   TS[126].ALLG.POS.End_1 := 491999;
   TS[126].ALLG.Stop_Position := 7200;
   TS[126].ALLG.Drive_speed_1 := 15000;
   TS[126].ALLG.Drive_speed_2 := 10000;
   TS[127].ALLG.POS.Start_1 := 492000;
   TS[127].ALLG.POS.End_1 := 498199;
   TS[127].ALLG.Stop_Position := 5400;
   TS[127].ALLG.Drive_speed_1 := 15000;
   TS[127].ALLG.Drive_speed_2 := 10000;
   TS[128].ALLG.POS.Start_1 := 498200;
   TS[128].ALLG.POS.End_1 := 504399;
   TS[128].ALLG.Stop_Position := 2954;
   TS[128].ALLG.Drive_speed_1 := 15000;
   TS[128].ALLG.Drive_speed_2 := 10000;
   TS[129].ALLG.POS.Start_1 := 504400;
   TS[129].ALLG.POS.End_1 := 511399;
   TS[129].ALLG.Stop_Position := 6300;
   TS[129].ALLG.Drive_speed_1 := 15000;
   TS[129].ALLG.Drive_speed_2 := 10000;
   TS[130].ALLG.POS.Start_1 := 511400;
   TS[130].ALLG.POS.End_1 := 518399;
   TS[130].ALLG.Stop_Position := 6300;
   TS[130].ALLG.Drive_speed_1 := 15000;
   TS[130].ALLG.Drive_speed_2 := 10000;
   TS[131].ALLG.POS.Start_1 := 518400;
   TS[131].ALLG.POS.End_1 := 525599;
   TS[131].ALLG.Stop_Position := 6300;
   TS[131].ALLG.Drive_speed_1 := 15000;
   TS[131].ALLG.Drive_speed_2 := 10000;
   TS[132].ALLG.POS.Start_1 := 525600;
   TS[132].ALLG.POS.End_1 := 529699;
   TS[132].ALLG.Stop_Position := 4299;
   TS[132].ALLG.Drive_speed_1 := 10000;
   TS[132].ALLG.Drive_speed_2 := 10000;
   TS[140].ALLG.POS.Start_1 := 529700;
   TS[140].ALLG.POS.End_1 := 535699;
   TS[140].ALLG.Stop_Position := 5900;
   TS[140].ALLG.Drive_speed_1 := 30000;
   TS[140].ALLG.Drive_speed_2 := 10000;
   TS[141].ALLG.POS.Start_1 := 535700;
   TS[141].ALLG.POS.End_1 := 541699;
   TS[141].ALLG.Stop_Position := 5900;
   TS[141].ALLG.Drive_speed_1 := 30000;
   TS[141].ALLG.Drive_speed_2 := 10000;
   TS[142].ALLG.POS.Start_1 := 541700;
   TS[142].ALLG.POS.End_1 := 547699;
   TS[142].ALLG.Stop_Position := 5900;
   TS[142].ALLG.Drive_speed_1 := 30000;
   TS[142].ALLG.Drive_speed_2 := 10000;
   TS[143].ALLG.POS.Start_1 := 547700;
   TS[143].ALLG.POS.End_1 := 553699;
   TS[143].ALLG.Stop_Position := 5900;
   TS[143].ALLG.Drive_speed_1 := 30000;
   TS[143].ALLG.Drive_speed_2 := 10000;
   TS[144].ALLG.POS.Start_1 := 553700;
   TS[144].ALLG.POS.End_1 := 559699;
   TS[144].ALLG.Stop_Position := 5900;
   TS[144].ALLG.Drive_speed_1 := 30000;
   TS[144].ALLG.Drive_speed_2 := 10000;
   TS[145].ALLG.POS.Start_1 := 559700;
   TS[145].ALLG.POS.End_1 := 565699;
   TS[145].ALLG.Stop_Position := 5900;
   TS[145].ALLG.Drive_speed_1 := 30000;
   TS[145].ALLG.Drive_speed_2 := 10000;
   TS[146].ALLG.POS.Start_1 := 565700;
   TS[146].ALLG.POS.End_1 := 571699;
   TS[146].ALLG.Stop_Position := 5900;
   TS[146].ALLG.Drive_speed_1 := 30000;
   TS[146].ALLG.Drive_speed_2 := 10000;
   TS[147].ALLG.POS.Start_1 := 571700;
   TS[147].ALLG.POS.End_1 := 577699;
   TS[147].ALLG.Stop_Position := 5900;
   TS[147].ALLG.Drive_speed_1 := 30000;
   TS[147].ALLG.Drive_speed_2 := 10000;
   TS[148].ALLG.POS.Start_1 := 577700;
   TS[148].ALLG.POS.End_1 := 583699;
   TS[148].ALLG.Stop_Position := 5900;
   TS[148].ALLG.Drive_speed_1 := 30000;
   TS[148].ALLG.Drive_speed_2 := 10000;
   TS[149].ALLG.POS.Start_1 := 583700;
   TS[149].ALLG.POS.End_1 := 589699;
   TS[149].ALLG.Stop_Position := 5900;
   TS[149].ALLG.Drive_speed_1 := 30000;
   TS[149].ALLG.Drive_speed_2 := 10000;
   TS[150].ALLG.POS.Start_1 := 589700;
   TS[150].ALLG.POS.End_1 := 595699;
   TS[150].ALLG.Stop_Position := 5900;
   TS[150].ALLG.Drive_speed_1 := 25000;
   TS[150].ALLG.Drive_speed_2 := 10000;
   TS[151].ALLG.POS.Start_1 := 595700;
   TS[151].ALLG.POS.End_1 := 601699;
   TS[151].ALLG.Stop_Position := 5900;
   TS[151].ALLG.Drive_speed_1 := 18000;
   TS[151].ALLG.Drive_speed_2 := 10000;
   TS[152].ALLG.POS.Start_1 := 601700;
   TS[152].ALLG.POS.End_1 := 607699;
   TS[152].ALLG.Stop_Position := 5900;
   TS[152].ALLG.Drive_speed_1 := 18000;
   TS[152].ALLG.Drive_speed_2 := 10000;
   TS[160].ALLG.POS.Start_1 := 607700;
   TS[160].ALLG.POS.End_1 := 613699;
   TS[160].ALLG.Stop_Position := 5900;
   TS[160].ALLG.Drive_speed_1 := 20000;
   TS[160].ALLG.Drive_speed_2 := 10000;
   TS[161].ALLG.POS.Start_1 := 613700;
   TS[161].ALLG.POS.End_1 := 619699;
   TS[161].ALLG.Stop_Position := 5900;
   TS[161].ALLG.Drive_speed_1 := 20000;
   TS[161].ALLG.Drive_speed_2 := 10000;
   TS[162].ALLG.POS.Start_1 := 619700;
   TS[162].ALLG.POS.End_1 := 625699;
   TS[162].ALLG.Stop_Position := 5900;
   TS[162].ALLG.Drive_speed_1 := 20000;
   TS[162].ALLG.Drive_speed_2 := 10000;
   // 15300 more start values not shown
END_DATA_BLOCK

DATA_BLOCK "DB_SDC_TS_PARAMETER_3"   // DB3706
{ S7_Optimized_Access := 'FALSE' }
AUTHOR : FFM
FAMILY : SDC
NAME : SECT_DEF
VERSION : 1.0
   VAR
      HEADER : Struct   // Struktur für Datenheader // nicht verschieben
         DB_NR : Int := 3706;   // DB Nummer
         MIN_NR_SEK : Int := 201;   // Niedrigste SEK Nummer im DB
         MAX_NR_SEK : Int := 300;   // Höchste SEK Nummer im DB
         START_DAT : Int := 20;   // Startadresse der SEK im DB
         LAENGE_SEK_DATA : Int := 260;   // Länge SEK Data
         ANZ_PROFIL : Int := 10;   // Number of Profiles
         OFFEST_PROFIL : Int := 40;   // Offestadresse der Profilparameter im TS-Parameterdatensatz
         LAENGE_PROFIL_DATA : Int := 22;   // Länge SEK Data
         Res160 : Int := 0;   // Reserve
         Res : Int := 0;   // Reserve
      END_STRUCT;
      TS : Array[201..300] of "UDT_SDC_TS_PARAMETER";
   END_VAR
BEGIN
   TS[201].ALLG.SEK_NEXT_1 := 0;
   TS[201].ALLG.SEK_NEXT_2 := 0;
   TS[201].ALLG.Spare[4] := 16#00;
   TS[201].ALLG.Spare[5] := 16#00;
   TS[201].ALLG.POS.Start_1 := 709550;
   TS[201].ALLG.POS.End_1 := 715849;
   TS[201].ALLG.POS.Start_2 := 0;
   TS[201].ALLG.POS.End_2 := 0;
   TS[201].ALLG.POS.Actionpoint_1 := 0;
   TS[201].ALLG.POS.Actionpoint_2 := 0;
   TS[201].ALLG.FLAGS.DIST_VAL[0] := FALSE;
   TS[201].ALLG.FLAGS.DIST_VAL[1] := FALSE;
   TS[201].ALLG.FLAGS.DIST_VAL[2] := FALSE;
   TS[201].ALLG.FLAGS.DIST_VAL[3] := FALSE;
   TS[201].ALLG.FLAGS.DIST_VAL[4] := FALSE;
   TS[201].ALLG.FLAGS.DIST_VAL[5] := FALSE;
   TS[201].ALLG.FLAGS.DIST_VAL[6] := FALSE;
   TS[201].ALLG.FLAGS.DIST_VAL[7] := FALSE;
   TS[201].ALLG.FLAGS.DIST_VAL[8] := FALSE;
   TS[201].ALLG.FLAGS.DIST_VAL[9] := TRUE;
   TS[201].ALLG.FLAGS.DIST_VAL[10] := FALSE;
   TS[201].ALLG.FLAGS.DIST_VAL[11] := FALSE;
   TS[201].ALLG.FLAGS.DIST_VAL[12] := FALSE;
   TS[201].ALLG.FLAGS.DIST_VAL[13] := FALSE;
   TS[201].ALLG.FLAGS.DIST_VAL[14] := FALSE;
   TS[201].ALLG.FLAGS.DIST_VAL[15] := FALSE;
   TS[201].ALLG.FLAGS.one_profile := FALSE;
   TS[201].ALLG.FLAGS.BLIND := FALSE;
   TS[201].ALLG.FLAGS.NO_DIST_CONT := FALSE;
   TS[201].ALLG.FLAGS.SYNCH_AREA := FALSE;
   TS[201].ALLG.FLAGS.bit24 := FALSE;
   TS[201].ALLG.FLAGS.bit25 := FALSE;
   TS[201].ALLG.FLAGS.bit26 := FALSE;
   TS[201].ALLG.FLAGS.bit27 := FALSE;
   TS[201].ALLG.FLAGS.EN_HOIST := FALSE;
   TS[201].ALLG.FLAGS.D_RESET_AFTER := FALSE;
   TS[201].ALLG.FLAGS.D_PULK := FALSE;
   TS[201].ALLG.FLAGS.bit33 := FALSE;
   TS[201].ALLG.FLAGS.bit34 := FALSE;
   TS[201].ALLG.FLAGS.bit35 := FALSE;
   TS[201].ALLG.FLAGS.bit36 := FALSE;
   TS[201].ALLG.FLAGS.Deutronic_ON := FALSE;
   TS[201].ALLG.Stop_Position := 5800;
   TS[201].ALLG.Drive_speed_1 := 18000;
   TS[201].ALLG.Drive_speed_2 := 6000;
   TS[201].PROFIL[1].Hoist_Pos_start := 0;
   TS[201].PROFIL[1].Height := 3890;
   TS[201].PROFIL[1].Hoist_speed := 2000;
   TS[201].PROFIL[1].Hoist_offset_1 := 0;
   TS[201].PROFIL[1].Hoist_offset_2 := 0;
   TS[201].PROFIL[1].Hoist_offset_3 := 0;
   TS[201].PROFIL[1].Hoist_offset_4 := 0;
   TS[201].PROFIL[1].Hoist_Start_offset_1 := 0;
   TS[201].PROFIL[1].Hoist_Start_offset_2 := 0;
   TS[201].PROFIL[1].Hoist_Start_offset_3 := 0;
   TS[201].PROFIL[1].Hoist_Start_offset_4 := 0;
   TS[201].PROFIL[2].Hoist_Pos_start := 0;
   TS[201].PROFIL[2].Height := 3890;
   TS[201].PROFIL[2].Hoist_speed := 2000;
   TS[201].PROFIL[2].Hoist_offset_1 := 0;
   TS[201].PROFIL[2].Hoist_offset_2 := 0;
   TS[201].PROFIL[2].Hoist_offset_3 := 0;
   TS[201].PROFIL[2].Hoist_offset_4 := 0;
   TS[201].PROFIL[2].Hoist_Start_offset_1 := 0;
   TS[201].PROFIL[2].Hoist_Start_offset_2 := 0;
   TS[201].PROFIL[2].Hoist_Start_offset_3 := 0;
   TS[201].PROFIL[2].Hoist_Start_offset_4 := 0;
   TS[201].PROFIL[3].Hoist_Pos_start := 0;
   TS[201].PROFIL[3].Height := 3890;
   TS[201].PROFIL[3].Hoist_speed := 2000;
   TS[201].PROFIL[3].Hoist_offset_1 := 0;
   TS[201].PROFIL[3].Hoist_offset_2 := 0;
   TS[201].PROFIL[3].Hoist_offset_3 := 0;
   TS[201].PROFIL[3].Hoist_offset_4 := 0;
   TS[201].PROFIL[3].Hoist_Start_offset_1 := 0;
   TS[201].PROFIL[3].Hoist_Start_offset_2 := 0;
   TS[201].PROFIL[3].Hoist_Start_offset_3 := 0;
   TS[201].PROFIL[3].Hoist_Start_offset_4 := 0;
   TS[201].PROFIL[4].Hoist_Pos_start := 0;
   TS[201].PROFIL[4].Height := 3890;
   TS[201].PROFIL[4].Hoist_speed := 2000;
   TS[201].PROFIL[4].Hoist_offset_1 := 0;
   TS[201].PROFIL[4].Hoist_offset_2 := 0;
   TS[201].PROFIL[4].Hoist_offset_3 := 0;
   TS[201].PROFIL[4].Hoist_offset_4 := 0;
   TS[201].PROFIL[4].Hoist_Start_offset_1 := 0;
   TS[201].PROFIL[4].Hoist_Start_offset_2 := 0;
   TS[201].PROFIL[4].Hoist_Start_offset_3 := 0;
   TS[201].PROFIL[4].Hoist_Start_offset_4 := 0;
   TS[201].PROFIL[5].Hoist_Pos_start := 0;
   TS[201].PROFIL[5].Height := 3890;
   TS[201].PROFIL[5].Hoist_speed := 2000;
   TS[201].PROFIL[5].Hoist_offset_1 := 0;
   TS[201].PROFIL[5].Hoist_offset_2 := 0;
   TS[201].PROFIL[5].Hoist_offset_3 := 0;
   TS[201].PROFIL[5].Hoist_offset_4 := 0;
   TS[201].PROFIL[5].Hoist_Start_offset_1 := 0;
   TS[201].PROFIL[5].Hoist_Start_offset_2 := 0;
   TS[201].PROFIL[5].Hoist_Start_offset_3 := 0;
   TS[201].PROFIL[5].Hoist_Start_offset_4 := 0;
   TS[201].PROFIL[6].Hoist_Pos_start := 0;
   TS[201].PROFIL[6].Height := 3890;
   TS[201].PROFIL[6].Hoist_speed := 2000;
   TS[201].PROFIL[6].Hoist_offset_1 := 0;
   TS[201].PROFIL[6].Hoist_offset_2 := 0;
   TS[201].PROFIL[6].Hoist_offset_3 := 0;
   TS[201].PROFIL[6].Hoist_offset_4 := 0;
   TS[201].PROFIL[6].Hoist_Start_offset_1 := 0;
   TS[201].PROFIL[6].Hoist_Start_offset_2 := 0;
   TS[201].PROFIL[6].Hoist_Start_offset_3 := 0;
   TS[201].PROFIL[6].Hoist_Start_offset_4 := 0;
   TS[201].PROFIL[7].Hoist_Pos_start := 0;
   TS[201].PROFIL[7].Height := 3890;
   TS[201].PROFIL[7].Hoist_speed := 2000;
   TS[201].PROFIL[7].Hoist_offset_1 := 0;
   TS[201].PROFIL[7].Hoist_offset_2 := 0;
   TS[201].PROFIL[7].Hoist_offset_3 := 0;
   TS[201].PROFIL[7].Hoist_offset_4 := 0;
   TS[201].PROFIL[7].Hoist_Start_offset_1 := 0;
   TS[201].PROFIL[7].Hoist_Start_offset_2 := 0;
   TS[201].PROFIL[7].Hoist_Start_offset_3 := 0;
   TS[201].PROFIL[7].Hoist_Start_offset_4 := 0;
   TS[201].PROFIL[8].Hoist_Pos_start := 0;
   TS[201].PROFIL[8].Height := 3890;
   TS[201].PROFIL[8].Hoist_speed := 2000;
   TS[201].PROFIL[8].Hoist_offset_1 := 0;
   TS[201].PROFIL[8].Hoist_offset_2 := 0;
   TS[201].PROFIL[8].Hoist_offset_3 := 0;
   TS[201].PROFIL[8].Hoist_offset_4 := 0;
   TS[201].PROFIL[8].Hoist_Start_offset_1 := 0;
   TS[201].PROFIL[8].Hoist_Start_offset_2 := 0;
   TS[201].PROFIL[8].Hoist_Start_offset_3 := 0;
   TS[201].PROFIL[8].Hoist_Start_offset_4 := 0;
   TS[201].PROFIL[9].Hoist_Pos_start := 0;
   TS[201].PROFIL[9].Height := 3890;
   TS[201].PROFIL[9].Hoist_speed := 2000;
   TS[201].PROFIL[9].Hoist_offset_1 := 0;
   TS[201].PROFIL[9].Hoist_offset_2 := 0;
   TS[201].PROFIL[9].Hoist_offset_3 := 0;
   TS[201].PROFIL[9].Hoist_offset_4 := 0;
   TS[201].PROFIL[9].Hoist_Start_offset_1 := 0;
   TS[201].PROFIL[9].Hoist_Start_offset_2 := 0;
   TS[201].PROFIL[9].Hoist_Start_offset_3 := 0;
   TS[201].PROFIL[9].Hoist_Start_offset_4 := 0;
   TS[201].PROFIL[10].Hoist_Pos_start := 0;
   TS[201].PROFIL[10].Height := 3890;
   TS[201].PROFIL[10].Hoist_speed := 2000;
   TS[201].PROFIL[10].Hoist_offset_1 := 0;
   TS[201].PROFIL[10].Hoist_offset_2 := 0;
   TS[201].PROFIL[10].Hoist_offset_3 := 0;
   TS[201].PROFIL[10].Hoist_offset_4 := 0;
   TS[201].PROFIL[10].Hoist_Start_offset_1 := 0;
   TS[201].PROFIL[10].Hoist_Start_offset_2 := 0;
   TS[201].PROFIL[10].Hoist_Start_offset_3 := 0;
   TS[201].PROFIL[10].Hoist_Start_offset_4 := 0;
   TS[202].ALLG.SEK_NEXT_1 := 0;
   TS[202].ALLG.SEK_NEXT_2 := 0;
   TS[202].ALLG.Spare[4] := 16#00;
   TS[202].ALLG.Spare[5] := 16#00;
   TS[202].ALLG.POS.Start_1 := 715850;
   TS[202].ALLG.POS.End_1 := 722149;
   TS[202].ALLG.POS.Start_2 := 0;
   TS[202].ALLG.POS.End_2 := 0;
   TS[202].ALLG.POS.Actionpoint_1 := 0;
   TS[202].ALLG.POS.Actionpoint_2 := 0;
   TS[202].ALLG.FLAGS.DIST_VAL[0] := FALSE;
   TS[202].ALLG.FLAGS.DIST_VAL[1] := FALSE;
   TS[202].ALLG.FLAGS.DIST_VAL[2] := FALSE;
   TS[202].ALLG.FLAGS.DIST_VAL[3] := FALSE;
   TS[202].ALLG.FLAGS.DIST_VAL[4] := FALSE;
   TS[202].ALLG.FLAGS.DIST_VAL[5] := FALSE;
   TS[202].ALLG.FLAGS.DIST_VAL[6] := FALSE;
   TS[202].ALLG.FLAGS.DIST_VAL[7] := FALSE;
   TS[202].ALLG.FLAGS.DIST_VAL[8] := FALSE;
   TS[202].ALLG.FLAGS.DIST_VAL[9] := TRUE;
   TS[202].ALLG.FLAGS.DIST_VAL[10] := FALSE;
   TS[202].ALLG.FLAGS.DIST_VAL[11] := FALSE;
   TS[202].ALLG.FLAGS.DIST_VAL[12] := FALSE;
   TS[202].ALLG.FLAGS.DIST_VAL[13] := FALSE;
   TS[202].ALLG.FLAGS.DIST_VAL[14] := FALSE;
   TS[202].ALLG.FLAGS.DIST_VAL[15] := FALSE;
   TS[202].ALLG.FLAGS.one_profile := FALSE;
   TS[202].ALLG.FLAGS.BLIND := FALSE;
   TS[202].ALLG.FLAGS.NO_DIST_CONT := FALSE;
   TS[202].ALLG.FLAGS.SYNCH_AREA := FALSE;
   TS[202].ALLG.FLAGS.bit24 := FALSE;
   TS[202].ALLG.FLAGS.bit25 := FALSE;
   TS[202].ALLG.FLAGS.bit26 := FALSE;
   TS[202].ALLG.FLAGS.bit27 := FALSE;
   TS[202].ALLG.FLAGS.EN_HOIST := FALSE;
   TS[202].ALLG.FLAGS.D_RESET_AFTER := FALSE;
   TS[202].ALLG.FLAGS.D_PULK := FALSE;
   TS[202].ALLG.FLAGS.bit33 := FALSE;
   TS[202].ALLG.FLAGS.bit34 := FALSE;
   TS[202].ALLG.FLAGS.bit35 := FALSE;
   TS[202].ALLG.FLAGS.bit36 := FALSE;
   TS[202].ALLG.FLAGS.Deutronic_ON := FALSE;
   TS[202].ALLG.Stop_Position := 5800;
   TS[202].ALLG.Drive_speed_1 := 18000;
   TS[202].ALLG.Drive_speed_2 := 6000;
   // 15300 more start values not shown
END_DATA_BLOCK

DATA_BLOCK "DB_SDC_TS_PARAMETER_4"   // DB3707
{ S7_Optimized_Access := 'FALSE' }
AUTHOR : FFM
FAMILY : SDC
NAME : SECT_DEF
VERSION : 1.0
   VAR
      HEADER : Struct   // Struktur für Datenheader // nicht verschieben
         DB_NR : Int := 3707;   // DB Nummer
         MIN_NR_SEK : Int := 301;   // Niedrigste SEK Nummer im DB
         MAX_NR_SEK : Int := 400;   // Höchste SEK Nummer im DB
         START_DAT : Int := 20;   // Startadresse der SEK im DB
         LAENGE_SEK_DATA : Int := 260;   // Länge SEK Data
         ANZ_PROFIL : Int := 10;   // Number of Profiles
         OFFEST_PROFIL : Int := 40;   // Offestadresse der Profilparameter im TS-Parameterdatensatz
         LAENGE_PROFIL_DATA : Int := 22;   // Länge SEK Data
         Res160 : Int := 0;   // Reserve
         Res : Int := 0;   // Reserve
      END_STRUCT;
      TS : Array[301..400] of "UDT_SDC_TS_PARAMETER";
   END_VAR
BEGIN
   TS[301].ALLG.SEK_NEXT_1 := 0;
   TS[301].ALLG.SEK_NEXT_2 := 0;
   TS[301].ALLG.Spare[4] := 16#00;
   TS[301].ALLG.Spare[5] := 16#00;
   TS[301].ALLG.POS.Start_1 := 0;
   TS[301].ALLG.POS.End_1 := 0;
   TS[301].ALLG.POS.Start_2 := 0;
   TS[301].ALLG.POS.End_2 := 0;
   TS[301].ALLG.POS.Actionpoint_1 := 0;
   TS[301].ALLG.POS.Actionpoint_2 := 0;
   TS[301].ALLG.FLAGS.DIST_VAL[0] := TRUE;
   TS[301].ALLG.FLAGS.DIST_VAL[1] := FALSE;
   TS[301].ALLG.FLAGS.DIST_VAL[2] := FALSE;
   TS[301].ALLG.FLAGS.DIST_VAL[3] := FALSE;
   TS[301].ALLG.FLAGS.DIST_VAL[4] := FALSE;
   TS[301].ALLG.FLAGS.DIST_VAL[5] := FALSE;
   TS[301].ALLG.FLAGS.DIST_VAL[6] := FALSE;
   TS[301].ALLG.FLAGS.DIST_VAL[7] := FALSE;
   TS[301].ALLG.FLAGS.DIST_VAL[8] := FALSE;
   TS[301].ALLG.FLAGS.DIST_VAL[9] := FALSE;
   TS[301].ALLG.FLAGS.DIST_VAL[10] := FALSE;
   TS[301].ALLG.FLAGS.DIST_VAL[11] := FALSE;
   TS[301].ALLG.FLAGS.DIST_VAL[12] := FALSE;
   TS[301].ALLG.FLAGS.DIST_VAL[13] := FALSE;
   TS[301].ALLG.FLAGS.DIST_VAL[14] := FALSE;
   TS[301].ALLG.FLAGS.DIST_VAL[15] := FALSE;
   TS[301].ALLG.FLAGS.one_profile := FALSE;
   TS[301].ALLG.FLAGS.BLIND := FALSE;
   TS[301].ALLG.FLAGS.NO_DIST_CONT := FALSE;
   TS[301].ALLG.FLAGS.SYNCH_AREA := FALSE;
   TS[301].ALLG.FLAGS.bit24 := FALSE;
   TS[301].ALLG.FLAGS.bit25 := FALSE;
   TS[301].ALLG.FLAGS.bit26 := FALSE;
   TS[301].ALLG.FLAGS.bit27 := FALSE;
   TS[301].ALLG.FLAGS.EN_HOIST := FALSE;
   TS[301].ALLG.FLAGS.D_RESET_AFTER := FALSE;
   TS[301].ALLG.FLAGS.D_PULK := FALSE;
   TS[301].ALLG.FLAGS.bit33 := FALSE;
   TS[301].ALLG.FLAGS.bit34 := FALSE;
   TS[301].ALLG.FLAGS.bit35 := FALSE;
   TS[301].ALLG.FLAGS.bit36 := FALSE;
   TS[301].ALLG.FLAGS.Deutronic_ON := FALSE;
   TS[301].ALLG.Stop_Position := 0;
   TS[301].ALLG.Drive_speed_1 := 0;
   TS[301].ALLG.Drive_speed_2 := 0;
   TS[301].PROFIL[1].Hoist_Pos_start := 0;
   TS[301].PROFIL[1].Height := 2651;
   TS[301].PROFIL[1].Hoist_speed := 2000;
   TS[301].PROFIL[1].Hoist_offset_1 := 0;
   TS[301].PROFIL[1].Hoist_offset_2 := 0;
   TS[301].PROFIL[1].Hoist_offset_3 := 0;
   TS[301].PROFIL[1].Hoist_offset_4 := 0;
   TS[301].PROFIL[1].Hoist_Start_offset_1 := 0;
   TS[301].PROFIL[1].Hoist_Start_offset_2 := 0;
   TS[301].PROFIL[1].Hoist_Start_offset_3 := 0;
   TS[301].PROFIL[1].Hoist_Start_offset_4 := 0;
   TS[301].PROFIL[2].Hoist_Pos_start := 0;
   TS[301].PROFIL[2].Height := 2651;
   TS[301].PROFIL[2].Hoist_speed := 2000;
   TS[301].PROFIL[2].Hoist_offset_1 := 0;
   TS[301].PROFIL[2].Hoist_offset_2 := 0;
   TS[301].PROFIL[2].Hoist_offset_3 := 0;
   TS[301].PROFIL[2].Hoist_offset_4 := 0;
   TS[301].PROFIL[2].Hoist_Start_offset_1 := 0;
   TS[301].PROFIL[2].Hoist_Start_offset_2 := 0;
   TS[301].PROFIL[2].Hoist_Start_offset_3 := 0;
   TS[301].PROFIL[2].Hoist_Start_offset_4 := 0;
   TS[301].PROFIL[3].Hoist_Pos_start := 0;
   TS[301].PROFIL[3].Height := 2651;
   TS[301].PROFIL[3].Hoist_speed := 2000;
   TS[301].PROFIL[3].Hoist_offset_1 := 0;
   TS[301].PROFIL[3].Hoist_offset_2 := 0;
   TS[301].PROFIL[3].Hoist_offset_3 := 0;
   TS[301].PROFIL[3].Hoist_offset_4 := 0;
   TS[301].PROFIL[3].Hoist_Start_offset_1 := 0;
   TS[301].PROFIL[3].Hoist_Start_offset_2 := 0;
   TS[301].PROFIL[3].Hoist_Start_offset_3 := 0;
   TS[301].PROFIL[3].Hoist_Start_offset_4 := 0;
   TS[301].PROFIL[4].Hoist_Pos_start := 0;
   TS[301].PROFIL[4].Height := 2651;
   TS[301].PROFIL[4].Hoist_speed := 2000;
   TS[301].PROFIL[4].Hoist_offset_1 := 0;
   TS[301].PROFIL[4].Hoist_offset_2 := 0;
   TS[301].PROFIL[4].Hoist_offset_3 := 0;
   TS[301].PROFIL[4].Hoist_offset_4 := 0;
   TS[301].PROFIL[4].Hoist_Start_offset_1 := 0;
   TS[301].PROFIL[4].Hoist_Start_offset_2 := 0;
   TS[301].PROFIL[4].Hoist_Start_offset_3 := 0;
   TS[301].PROFIL[4].Hoist_Start_offset_4 := 0;
   TS[301].PROFIL[5].Hoist_Pos_start := 0;
   TS[301].PROFIL[5].Height := 2651;
   TS[301].PROFIL[5].Hoist_speed := 2000;
   TS[301].PROFIL[5].Hoist_offset_1 := 0;
   TS[301].PROFIL[5].Hoist_offset_2 := 0;
   TS[301].PROFIL[5].Hoist_offset_3 := 0;
   TS[301].PROFIL[5].Hoist_offset_4 := 0;
   TS[301].PROFIL[5].Hoist_Start_offset_1 := 0;
   TS[301].PROFIL[5].Hoist_Start_offset_2 := 0;
   TS[301].PROFIL[5].Hoist_Start_offset_3 := 0;
   TS[301].PROFIL[5].Hoist_Start_offset_4 := 0;
   TS[301].PROFIL[6].Hoist_Pos_start := 0;
   TS[301].PROFIL[6].Height := 2651;
   TS[301].PROFIL[6].Hoist_speed := 2000;
   TS[301].PROFIL[6].Hoist_offset_1 := 0;
   TS[301].PROFIL[6].Hoist_offset_2 := 0;
   TS[301].PROFIL[6].Hoist_offset_3 := 0;
   TS[301].PROFIL[6].Hoist_offset_4 := 0;
   TS[301].PROFIL[6].Hoist_Start_offset_1 := 0;
   TS[301].PROFIL[6].Hoist_Start_offset_2 := 0;
   TS[301].PROFIL[6].Hoist_Start_offset_3 := 0;
   TS[301].PROFIL[6].Hoist_Start_offset_4 := 0;
   TS[301].PROFIL[7].Hoist_Pos_start := 0;
   TS[301].PROFIL[7].Height := 2651;
   TS[301].PROFIL[7].Hoist_speed := 2000;
   TS[301].PROFIL[7].Hoist_offset_1 := 0;
   TS[301].PROFIL[7].Hoist_offset_2 := 0;
   TS[301].PROFIL[7].Hoist_offset_3 := 0;
   TS[301].PROFIL[7].Hoist_offset_4 := 0;
   TS[301].PROFIL[7].Hoist_Start_offset_1 := 0;
   TS[301].PROFIL[7].Hoist_Start_offset_2 := 0;
   TS[301].PROFIL[7].Hoist_Start_offset_3 := 0;
   TS[301].PROFIL[7].Hoist_Start_offset_4 := 0;
   TS[301].PROFIL[8].Hoist_Pos_start := 0;
   TS[301].PROFIL[8].Height := 2651;
   TS[301].PROFIL[8].Hoist_speed := 2000;
   TS[301].PROFIL[8].Hoist_offset_1 := 0;
   TS[301].PROFIL[8].Hoist_offset_2 := 0;
   TS[301].PROFIL[8].Hoist_offset_3 := 0;
   TS[301].PROFIL[8].Hoist_offset_4 := 0;
   TS[301].PROFIL[8].Hoist_Start_offset_1 := 0;
   TS[301].PROFIL[8].Hoist_Start_offset_2 := 0;
   TS[301].PROFIL[8].Hoist_Start_offset_3 := 0;
   TS[301].PROFIL[8].Hoist_Start_offset_4 := 0;
   TS[301].PROFIL[9].Hoist_Pos_start := 0;
   TS[301].PROFIL[9].Height := 2651;
   TS[301].PROFIL[9].Hoist_speed := 2000;
   TS[301].PROFIL[9].Hoist_offset_1 := 0;
   TS[301].PROFIL[9].Hoist_offset_2 := 0;
   TS[301].PROFIL[9].Hoist_offset_3 := 0;
   TS[301].PROFIL[9].Hoist_offset_4 := 0;
   TS[301].PROFIL[9].Hoist_Start_offset_1 := 0;
   TS[301].PROFIL[9].Hoist_Start_offset_2 := 0;
   TS[301].PROFIL[9].Hoist_Start_offset_3 := 0;
   TS[301].PROFIL[9].Hoist_Start_offset_4 := 0;
   TS[301].PROFIL[10].Hoist_Pos_start := 0;
   TS[301].PROFIL[10].Height := 2651;
   TS[301].PROFIL[10].Hoist_speed := 2000;
   TS[301].PROFIL[10].Hoist_offset_1 := 0;
   TS[301].PROFIL[10].Hoist_offset_2 := 0;
   TS[301].PROFIL[10].Hoist_offset_3 := 0;
   TS[301].PROFIL[10].Hoist_offset_4 := 0;
   TS[301].PROFIL[10].Hoist_Start_offset_1 := 0;
   TS[301].PROFIL[10].Hoist_Start_offset_2 := 0;
   TS[301].PROFIL[10].Hoist_Start_offset_3 := 0;
   TS[301].PROFIL[10].Hoist_Start_offset_4 := 0;
   TS[302].ALLG.SEK_NEXT_1 := 0;
   TS[302].ALLG.SEK_NEXT_2 := 0;
   TS[302].ALLG.Spare[4] := 16#00;
   TS[302].ALLG.Spare[5] := 16#00;
   TS[302].ALLG.POS.Start_1 := 0;
   TS[302].ALLG.POS.End_1 := 0;
   TS[302].ALLG.POS.Start_2 := 0;
   TS[302].ALLG.POS.End_2 := 0;
   TS[302].ALLG.POS.Actionpoint_1 := 0;
   TS[302].ALLG.POS.Actionpoint_2 := 0;
   TS[302].ALLG.FLAGS.DIST_VAL[0] := TRUE;
   TS[302].ALLG.FLAGS.DIST_VAL[1] := FALSE;
   TS[302].ALLG.FLAGS.DIST_VAL[2] := FALSE;
   TS[302].ALLG.FLAGS.DIST_VAL[3] := FALSE;
   TS[302].ALLG.FLAGS.DIST_VAL[4] := FALSE;
   TS[302].ALLG.FLAGS.DIST_VAL[5] := FALSE;
   TS[302].ALLG.FLAGS.DIST_VAL[6] := FALSE;
   TS[302].ALLG.FLAGS.DIST_VAL[7] := FALSE;
   TS[302].ALLG.FLAGS.DIST_VAL[8] := FALSE;
   TS[302].ALLG.FLAGS.DIST_VAL[9] := FALSE;
   TS[302].ALLG.FLAGS.DIST_VAL[10] := FALSE;
   TS[302].ALLG.FLAGS.DIST_VAL[11] := FALSE;
   TS[302].ALLG.FLAGS.DIST_VAL[12] := FALSE;
   TS[302].ALLG.FLAGS.DIST_VAL[13] := FALSE;
   TS[302].ALLG.FLAGS.DIST_VAL[14] := FALSE;
   TS[302].ALLG.FLAGS.DIST_VAL[15] := FALSE;
   TS[302].ALLG.FLAGS.one_profile := FALSE;
   TS[302].ALLG.FLAGS.BLIND := FALSE;
   TS[302].ALLG.FLAGS.NO_DIST_CONT := FALSE;
   TS[302].ALLG.FLAGS.SYNCH_AREA := FALSE;
   TS[302].ALLG.FLAGS.bit24 := FALSE;
   TS[302].ALLG.FLAGS.bit25 := FALSE;
   TS[302].ALLG.FLAGS.bit26 := FALSE;
   TS[302].ALLG.FLAGS.bit27 := FALSE;
   TS[302].ALLG.FLAGS.EN_HOIST := FALSE;
   TS[302].ALLG.FLAGS.D_RESET_AFTER := FALSE;
   TS[302].ALLG.FLAGS.D_PULK := FALSE;
   TS[302].ALLG.FLAGS.bit33 := FALSE;
   TS[302].ALLG.FLAGS.bit34 := FALSE;
   TS[302].ALLG.FLAGS.bit35 := FALSE;
   TS[302].ALLG.FLAGS.bit36 := FALSE;
   TS[302].ALLG.FLAGS.Deutronic_ON := FALSE;
   TS[302].ALLG.Stop_Position := 0;
   TS[302].ALLG.Drive_speed_1 := 0;
   TS[302].ALLG.Drive_speed_2 := 0;
   // 15300 more start values not shown
END_DATA_BLOCK

DATA_BLOCK "DB_SDC_TS_PARAMETER_5"   // DB3708
{ S7_Optimized_Access := 'FALSE' }
AUTHOR : FFM
FAMILY : SDC
NAME : SECT_DEF
VERSION : 1.0
   VAR
      HEADER : Struct   // Struktur für Datenheader // nicht verschieben
         DB_NR : Int := 3708;   // DB Nummer
         MIN_NR_SEK : Int := 401;   // Niedrigste SEK Nummer im DB
         MAX_NR_SEK : Int := 500;   // Höchste SEK Nummer im DB
         START_DAT : Int := 20;   // Startadresse der SEK im DB
         LAENGE_SEK_DATA : Int := 260;   // Länge SEK Data
         ANZ_PROFIL : Int := 10;   // Number of Profiles
         OFFEST_PROFIL : Int := 40;   // Offestadresse der Profilparameter im TS-Parameterdatensatz
         LAENGE_PROFIL_DATA : Int := 22;   // Länge SEK Data
         Res160 : Int := 0;   // Reserve
         Res : Int := 0;   // Reserve
      END_STRUCT;
      TS : Array[401..500] of "UDT_SDC_TS_PARAMETER";
   END_VAR
BEGIN
   TS[401].ALLG.SEK_NEXT_1 := 0;
   TS[401].ALLG.SEK_NEXT_2 := 0;
   TS[401].ALLG.Spare[4] := 16#00;
   TS[401].ALLG.Spare[5] := 16#00;
   TS[401].ALLG.POS.Start_1 := 1159500;
   TS[401].ALLG.POS.End_1 := 1165999;
   TS[401].ALLG.POS.Start_2 := 0;
   TS[401].ALLG.POS.End_2 := 0;
   TS[401].ALLG.POS.Actionpoint_1 := 0;
   TS[401].ALLG.POS.Actionpoint_2 := 0;
   TS[401].ALLG.FLAGS.DIST_VAL[0] := FALSE;
   TS[401].ALLG.FLAGS.DIST_VAL[1] := FALSE;
   TS[401].ALLG.FLAGS.DIST_VAL[2] := FALSE;
   TS[401].ALLG.FLAGS.DIST_VAL[3] := FALSE;
   TS[401].ALLG.FLAGS.DIST_VAL[4] := FALSE;
   TS[401].ALLG.FLAGS.DIST_VAL[5] := FALSE;
   TS[401].ALLG.FLAGS.DIST_VAL[6] := FALSE;
   TS[401].ALLG.FLAGS.DIST_VAL[7] := FALSE;
   TS[401].ALLG.FLAGS.DIST_VAL[8] := FALSE;
   TS[401].ALLG.FLAGS.DIST_VAL[9] := TRUE;
   TS[401].ALLG.FLAGS.DIST_VAL[10] := FALSE;
   TS[401].ALLG.FLAGS.DIST_VAL[11] := FALSE;
   TS[401].ALLG.FLAGS.DIST_VAL[12] := FALSE;
   TS[401].ALLG.FLAGS.DIST_VAL[13] := FALSE;
   TS[401].ALLG.FLAGS.DIST_VAL[14] := FALSE;
   TS[401].ALLG.FLAGS.DIST_VAL[15] := FALSE;
   TS[401].ALLG.FLAGS.one_profile := FALSE;
   TS[401].ALLG.FLAGS.BLIND := FALSE;
   TS[401].ALLG.FLAGS.NO_DIST_CONT := FALSE;
   TS[401].ALLG.FLAGS.SYNCH_AREA := FALSE;
   TS[401].ALLG.FLAGS.bit24 := FALSE;
   TS[401].ALLG.FLAGS.bit25 := FALSE;
   TS[401].ALLG.FLAGS.bit26 := FALSE;
   TS[401].ALLG.FLAGS.bit27 := FALSE;
   TS[401].ALLG.FLAGS.EN_HOIST := FALSE;
   TS[401].ALLG.FLAGS.D_RESET_AFTER := FALSE;
   TS[401].ALLG.FLAGS.D_PULK := FALSE;
   TS[401].ALLG.FLAGS.bit33 := FALSE;
   TS[401].ALLG.FLAGS.bit34 := FALSE;
   TS[401].ALLG.FLAGS.bit35 := FALSE;
   TS[401].ALLG.FLAGS.bit36 := FALSE;
   TS[401].ALLG.FLAGS.Deutronic_ON := FALSE;
   TS[401].ALLG.Stop_Position := 5800;
   TS[401].ALLG.Drive_speed_1 := 15000;
   TS[401].ALLG.Drive_speed_2 := 6000;
   TS[401].PROFIL[1].Hoist_Pos_start := 0;
   TS[401].PROFIL[1].Height := 3890;
   TS[401].PROFIL[1].Hoist_speed := 2000;
   TS[401].PROFIL[1].Hoist_offset_1 := 0;
   TS[401].PROFIL[1].Hoist_offset_2 := 0;
   TS[401].PROFIL[1].Hoist_offset_3 := 0;
   TS[401].PROFIL[1].Hoist_offset_4 := 0;
   TS[401].PROFIL[1].Hoist_Start_offset_1 := 0;
   TS[401].PROFIL[1].Hoist_Start_offset_2 := 0;
   TS[401].PROFIL[1].Hoist_Start_offset_3 := 0;
   TS[401].PROFIL[1].Hoist_Start_offset_4 := 0;
   TS[401].PROFIL[2].Hoist_Pos_start := 0;
   TS[401].PROFIL[2].Height := 3890;
   TS[401].PROFIL[2].Hoist_speed := 2000;
   TS[401].PROFIL[2].Hoist_offset_1 := 0;
   TS[401].PROFIL[2].Hoist_offset_2 := 0;
   TS[401].PROFIL[2].Hoist_offset_3 := 0;
   TS[401].PROFIL[2].Hoist_offset_4 := 0;
   TS[401].PROFIL[2].Hoist_Start_offset_1 := 0;
   TS[401].PROFIL[2].Hoist_Start_offset_2 := 0;
   TS[401].PROFIL[2].Hoist_Start_offset_3 := 0;
   TS[401].PROFIL[2].Hoist_Start_offset_4 := 0;
   TS[401].PROFIL[3].Hoist_Pos_start := 0;
   TS[401].PROFIL[3].Height := 3890;
   TS[401].PROFIL[3].Hoist_speed := 2000;
   TS[401].PROFIL[3].Hoist_offset_1 := 0;
   TS[401].PROFIL[3].Hoist_offset_2 := 0;
   TS[401].PROFIL[3].Hoist_offset_3 := 0;
   TS[401].PROFIL[3].Hoist_offset_4 := 0;
   TS[401].PROFIL[3].Hoist_Start_offset_1 := 0;
   TS[401].PROFIL[3].Hoist_Start_offset_2 := 0;
   TS[401].PROFIL[3].Hoist_Start_offset_3 := 0;
   TS[401].PROFIL[3].Hoist_Start_offset_4 := 0;
   TS[401].PROFIL[4].Hoist_Pos_start := 0;
   TS[401].PROFIL[4].Height := 3890;
   TS[401].PROFIL[4].Hoist_speed := 2000;
   TS[401].PROFIL[4].Hoist_offset_1 := 0;
   TS[401].PROFIL[4].Hoist_offset_2 := 0;
   TS[401].PROFIL[4].Hoist_offset_3 := 0;
   TS[401].PROFIL[4].Hoist_offset_4 := 0;
   TS[401].PROFIL[4].Hoist_Start_offset_1 := 0;
   TS[401].PROFIL[4].Hoist_Start_offset_2 := 0;
   TS[401].PROFIL[4].Hoist_Start_offset_3 := 0;
   TS[401].PROFIL[4].Hoist_Start_offset_4 := 0;
   TS[401].PROFIL[5].Hoist_Pos_start := 0;
   TS[401].PROFIL[5].Height := 3890;
   TS[401].PROFIL[5].Hoist_speed := 2000;
   TS[401].PROFIL[5].Hoist_offset_1 := 0;
   TS[401].PROFIL[5].Hoist_offset_2 := 0;
   TS[401].PROFIL[5].Hoist_offset_3 := 0;
   TS[401].PROFIL[5].Hoist_offset_4 := 0;
   TS[401].PROFIL[5].Hoist_Start_offset_1 := 0;
   TS[401].PROFIL[5].Hoist_Start_offset_2 := 0;
   TS[401].PROFIL[5].Hoist_Start_offset_3 := 0;
   TS[401].PROFIL[5].Hoist_Start_offset_4 := 0;
   TS[401].PROFIL[6].Hoist_Pos_start := 0;
   TS[401].PROFIL[6].Height := 3890;
   TS[401].PROFIL[6].Hoist_speed := 2000;
   TS[401].PROFIL[6].Hoist_offset_1 := 0;
   TS[401].PROFIL[6].Hoist_offset_2 := 0;
   TS[401].PROFIL[6].Hoist_offset_3 := 0;
   TS[401].PROFIL[6].Hoist_offset_4 := 0;
   TS[401].PROFIL[6].Hoist_Start_offset_1 := 0;
   TS[401].PROFIL[6].Hoist_Start_offset_2 := 0;
   TS[401].PROFIL[6].Hoist_Start_offset_3 := 0;
   TS[401].PROFIL[6].Hoist_Start_offset_4 := 0;
   TS[401].PROFIL[7].Hoist_Pos_start := 0;
   TS[401].PROFIL[7].Height := 3890;
   TS[401].PROFIL[7].Hoist_speed := 2000;
   TS[401].PROFIL[7].Hoist_offset_1 := 0;
   TS[401].PROFIL[7].Hoist_offset_2 := 0;
   TS[401].PROFIL[7].Hoist_offset_3 := 0;
   TS[401].PROFIL[7].Hoist_offset_4 := 0;
   TS[401].PROFIL[7].Hoist_Start_offset_1 := 0;
   TS[401].PROFIL[7].Hoist_Start_offset_2 := 0;
   TS[401].PROFIL[7].Hoist_Start_offset_3 := 0;
   TS[401].PROFIL[7].Hoist_Start_offset_4 := 0;
   TS[401].PROFIL[8].Hoist_Pos_start := 0;
   TS[401].PROFIL[8].Height := 3890;
   TS[401].PROFIL[8].Hoist_speed := 2000;
   TS[401].PROFIL[8].Hoist_offset_1 := 0;
   TS[401].PROFIL[8].Hoist_offset_2 := 0;
   TS[401].PROFIL[8].Hoist_offset_3 := 0;
   TS[401].PROFIL[8].Hoist_offset_4 := 0;
   TS[401].PROFIL[8].Hoist_Start_offset_1 := 0;
   TS[401].PROFIL[8].Hoist_Start_offset_2 := 0;
   TS[401].PROFIL[8].Hoist_Start_offset_3 := 0;
   TS[401].PROFIL[8].Hoist_Start_offset_4 := 0;
   TS[401].PROFIL[9].Hoist_Pos_start := 0;
   TS[401].PROFIL[9].Height := 3890;
   TS[401].PROFIL[9].Hoist_speed := 2000;
   TS[401].PROFIL[9].Hoist_offset_1 := 0;
   TS[401].PROFIL[9].Hoist_offset_2 := 0;
   TS[401].PROFIL[9].Hoist_offset_3 := 0;
   TS[401].PROFIL[9].Hoist_offset_4 := 0;
   TS[401].PROFIL[9].Hoist_Start_offset_1 := 0;
   TS[401].PROFIL[9].Hoist_Start_offset_2 := 0;
   TS[401].PROFIL[9].Hoist_Start_offset_3 := 0;
   TS[401].PROFIL[9].Hoist_Start_offset_4 := 0;
   TS[401].PROFIL[10].Hoist_Pos_start := 0;
   TS[401].PROFIL[10].Height := 3890;
   TS[401].PROFIL[10].Hoist_speed := 2000;
   TS[401].PROFIL[10].Hoist_offset_1 := 0;
   TS[401].PROFIL[10].Hoist_offset_2 := 0;
   TS[401].PROFIL[10].Hoist_offset_3 := 0;
   TS[401].PROFIL[10].Hoist_offset_4 := 0;
   TS[401].PROFIL[10].Hoist_Start_offset_1 := 0;
   TS[401].PROFIL[10].Hoist_Start_offset_2 := 0;
   TS[401].PROFIL[10].Hoist_Start_offset_3 := 0;
   TS[401].PROFIL[10].Hoist_Start_offset_4 := 0;
   TS[402].ALLG.SEK_NEXT_1 := 0;
   TS[402].ALLG.SEK_NEXT_2 := 0;
   TS[402].ALLG.Spare[4] := 16#00;
   TS[402].ALLG.Spare[5] := 16#00;
   TS[402].ALLG.POS.Start_1 := 1166000;
   TS[402].ALLG.POS.End_1 := 1172199;
   TS[402].ALLG.POS.Start_2 := 0;
   TS[402].ALLG.POS.End_2 := 0;
   TS[402].ALLG.POS.Actionpoint_1 := 0;
   TS[402].ALLG.POS.Actionpoint_2 := 0;
   TS[402].ALLG.FLAGS.DIST_VAL[0] := FALSE;
   TS[402].ALLG.FLAGS.DIST_VAL[1] := FALSE;
   TS[402].ALLG.FLAGS.DIST_VAL[2] := FALSE;
   TS[402].ALLG.FLAGS.DIST_VAL[3] := FALSE;
   TS[402].ALLG.FLAGS.DIST_VAL[4] := FALSE;
   TS[402].ALLG.FLAGS.DIST_VAL[5] := TRUE;
   TS[402].ALLG.FLAGS.DIST_VAL[6] := FALSE;
   TS[402].ALLG.FLAGS.DIST_VAL[7] := FALSE;
   TS[402].ALLG.FLAGS.DIST_VAL[8] := FALSE;
   TS[402].ALLG.FLAGS.DIST_VAL[9] := FALSE;
   TS[402].ALLG.FLAGS.DIST_VAL[10] := FALSE;
   TS[402].ALLG.FLAGS.DIST_VAL[11] := FALSE;
   TS[402].ALLG.FLAGS.DIST_VAL[12] := FALSE;
   TS[402].ALLG.FLAGS.DIST_VAL[13] := FALSE;
   TS[402].ALLG.FLAGS.DIST_VAL[14] := FALSE;
   TS[402].ALLG.FLAGS.DIST_VAL[15] := FALSE;
   TS[402].ALLG.FLAGS.one_profile := FALSE;
   TS[402].ALLG.FLAGS.BLIND := FALSE;
   TS[402].ALLG.FLAGS.NO_DIST_CONT := FALSE;
   TS[402].ALLG.FLAGS.SYNCH_AREA := FALSE;
   TS[402].ALLG.FLAGS.bit24 := FALSE;
   TS[402].ALLG.FLAGS.bit25 := FALSE;
   TS[402].ALLG.FLAGS.bit26 := FALSE;
   TS[402].ALLG.FLAGS.bit27 := FALSE;
   TS[402].ALLG.FLAGS.EN_HOIST := FALSE;
   TS[402].ALLG.FLAGS.D_RESET_AFTER := FALSE;
   TS[402].ALLG.FLAGS.D_PULK := FALSE;
   TS[402].ALLG.FLAGS.bit33 := FALSE;
   TS[402].ALLG.FLAGS.bit34 := FALSE;
   TS[402].ALLG.FLAGS.bit35 := FALSE;
   TS[402].ALLG.FLAGS.bit36 := FALSE;
   TS[402].ALLG.FLAGS.Deutronic_ON := FALSE;
   TS[402].ALLG.Stop_Position := 5800;
   TS[402].ALLG.Drive_speed_1 := 15000;
   TS[402].ALLG.Drive_speed_2 := 6000;
   // 15300 more start values not shown
END_DATA_BLOCK

